		
		2:(*//料框位置抓取*)		
		IF ii=129 THEN(*129表示所有有问题的都抓完了*)
			m_iStep:=4;
		ELSIF ii>0 AND ii<129 AND m_iCheck<>0 
					AND NOT FanucRobotIO.i_xBatteryDetect[0]
					AND NOT FanucRobotIO.i_xBatteryDetect[1]
					AND NOT FanucRobotIO.i_xBatteryDetect[2]
					AND NOT FanucRobotIO.i_xBatteryDetect[3](*4个电池位没料*)
					 (*有不良品*)THEN
			FanucRobotIO.o_xSortStart:=1;(*//从料框取料*)
			FanucRobotIO.o_xColumn[3]:=m_iCoordinateX/8=1;(*XY的偏移量计算在末尾*)
			FanucRobotIO.o_xColumn[2]:=(m_iCoordinateX MOD 8)/4=1;
			FanucRobotIO.o_xColumn[1]:=(m_iCoordinateX MOD 4)/2=1;
			FanucRobotIO.o_xColumn[0]:=(m_iCoordinateX MOD 2)/1=1;
			FanucRobotIO.o_xRow[3]:=m_iCoordinateY/8=1;			
			FanucRobotIO.o_xRow[2]:=(m_iCoordinateY MOD 8)/4=1;
			FanucRobotIO.o_xRow[1]:=(m_iCoordinateY MOD 4)/2=1;
			FanucRobotIO.o_xRow[0]:=(m_iCoordinateY MOD 2)/1=1;
			CASE SortCommunicationIO.i_arriBatteryStatus[ii] OF
			0:(*0表示OCV2的不良品，视为阻值错误处理*)
					FanucRobotIO.o_xPutNumber[1]:=1;					
			1:(*合格*)
					;
			2:(*容量不足*)
					FanucRobotIO.o_xPutNumber[0]:=1;	
			3:(*电压不足*)
					FanucRobotIO.o_xPutNumber[1]:=1;	
			4:(*阻值错误*)
					FanucRobotIO.o_xPutNumber[2]:=1;	
			5:(*电压过高*)
					FanucRobotIO.o_xPutNumber[3]:=1;	
			END_CASE;
		END_IF;
		IF FanucRobotIO.i_xPickOver THEN(*//抓取动作完成*)
			m_iStep:=3;
		END_IF;
	
		3:(*//放入下料皮带线*)
			FanucRobotIO.o_xSortStart:=0;(*//从料框取料*)
			FanucRobotIO.o_xColumn[3]:=0;(*XY的偏移量计算在末尾*)
			FanucRobotIO.o_xColumn[2]:=0;
			FanucRobotIO.o_xColumn[1]:=0;
			FanucRobotIO.o_xColumn[0]:=0;
			FanucRobotIO.o_xRow[3]:=0;
			FanucRobotIO.o_xRow[2]:=0;
			FanucRobotIO.o_xRow[1]:=0;
			FanucRobotIO.o_xRow[0]:=0;	
		IF FanucRobotIO.i_xPutOver THEN(*//抓取动作完成*)
			(*这个得放货完成在复位，方便step2给*)
			FanucRobotIO.o_xPutNumber[0]:=0;
			FanucRobotIO.o_xPutNumber[1]:=0;
			FanucRobotIO.o_xPutNumber[2]:=0;
			FanucRobotIO.o_xPutNumber[3]:=0;
		END_IF;
		m_TONPutover(IN:= FanucRobotIO.o_xPutNumber[0]=0
												AND FanucRobotIO.o_xPutNumber[1]=0
												AND FanucRobotIO.o_xPutNumber[2]=0
												AND FanucRobotIO.o_xPutNumber[3]=0,
			PT:=t#100ms ,Q:= m_xPutover,ET:=m_tPutover );	
			IF LDp(TRUE,m_xPutover)  THEN
				m_iStep:=2;
			END_IF;

		
		4:
		(*4复位所有数据*)
			FanucRobotIO.o_xSortStart:=0;(*//从料框取料*)
			FanucRobotIO.o_xColumn[3]:=0;(*XY的偏移量计算在末尾*)
			FanucRobotIO.o_xColumn[2]:=0;
			FanucRobotIO.o_xColumn[1]:=0;
			FanucRobotIO.o_xColumn[0]:=0;
			FanucRobotIO.o_xRow[3]:=0;
			FanucRobotIO.o_xRow[2]:=0;
			FanucRobotIO.o_xRow[1]:=0;
			FanucRobotIO.o_xRow[0]:=0;	
			FanucRobotIO.o_xPutNumber[0]:=0;
			FanucRobotIO.o_xPutNumber[1]:=0;
			FanucRobotIO.o_xPutNumber[2]:=0;
			FanucRobotIO.o_xPutNumber[3]:=0;

		IF  NOT SortCommunicationIO.o_xSortDone  THEN(*这里表示只给一下2*)
				SortCommunicationIO.o_iSortDonePLCPC:=2;
				SortCommunicationIO.o_xSortDone:=1;
		END_IF;		
		IF SortCommunicationIO.i_iSortDoneAknPCPLC =2 THEN
			SortCommunicationIO.o_iSortDonePLCPC:=1;
			m_iCoordinateX:=1;
			m_iCoordinateY:=1;
		END_IF;
	END_CASE;			
		IF ConveyorIO.xEmpty THEN
				m_iStep:=0;
		END_IF;

	m_iCheck:=	SortCommunicationIO.i_arriBatteryStatus[5]+
							SortCommunicationIO.i_arriBatteryStatus[1]+
							SortCommunicationIO.i_arriBatteryStatus[2]+
							SortCommunicationIO.i_arriBatteryStatus[3]+
							SortCommunicationIO.i_arriBatteryStatus[4];(*连续5个电池都是0，说明这框电池没数据，就不分拣*)
	IF LDP(TRUE,m_iStep=2 AND SortCommunicationIO.i_iInfoWriteDone=2 AND m_iCheck<>0) THEN(*判断哪个地方是有问题的*)
		FOR ii:=ii+1 TO 128 BY 1 DO
			IF SortCommunicationIO.i_arriBatteryStatus[ii]<>1 AND SortCommunicationIO.i_arriBatteryStatus[ii]<>5THEN
				m_iCoordinateX:=((ii-1)/ROW_NUB);
				m_iCoordinateY:=2*((ii-1)MOD ROW_NUB)+((m_iCoordinateX+1) MOD 2);(*把上位机给的编号值对应到二维的偏移上*)(*后面这个意思奇数排+1，偶数排不加*)
				EXIT;
			END_IF;
		END_FOR;
	END_IF;
END_IF;(*g_xauto*)	
IF  g_diDeviceIDSelect=ConveyorIO.diDeviceID AND g_xResetSingle THEN(*复位线体时，同时复位步数和请求，重新来一遍*)
	m_iStep:=0;
END_IF;	
IF  NOT g_xAuto THEN
		SortCommunicationIO.o_iRequestPLCPC:=0;
		SortCommunicationIO.o_iSortDonePLCPC:=0;
END_IF;
END_FUNCTION_BLOCK

PROGRAM START
IF g_xReset THEN
	SM50:=1;
	ELSE
	SM50:=0;
END_IF;
CASE g_iState OF
	0: (*手动*)
	g_xManual:=1;
	g_xAuto:=0;	
	g_xStackLampAmber:=1;
	g_xStackLampGreen:=0;
	g_xRemoteAuto:=0;
	g_xAutoLamp:=0;
	1:(*自动*)
	g_xManual:=0;
	g_xAuto:=1;
	g_xStackLampGreen:=1;
	g_xStackLampAmber:=0;
	g_xRemoteAuto:=0;
	g_xAutoLamp:=1;
	2:	(*远程自动*)
	g_xRemoteAuto:=1;
	g_xStackLampGreen:=1;
	g_xStackLampAmber:=0;
	g_xAuto:=0;
	g_xManual:=0;
	g_xAutoLamp:=0;
	3:(*自动未启动*)
	g_xRemoteAuto:=1;
	g_xStackLampGreen:=SM412;
	g_xStackLampAmber:=0;
	g_xAuto:=0;
	g_xManual:=0;	
	g_xAutoLamp:=0;
END_CASE;

IF g_xAutoSwitch AND g_xAutoStart  THEN  
	g_iState:=1;
END_IF;

IF g_xAutoSwitch AND (g_iState<>1 OR NOT g_xStop)  THEN  
	g_iState:=3;
END_IF;

g_xStackLampRed:=g_xAlarm AND SM412;
g_xBuzzer:=g_xAlarm AND SM412 AND NOT g_xMute;

IF LDF(TRUE,g_xAlarm) THEN
	g_xMute:=0;
END_IF;

IF NOT g_xAutoSwitch  OR g_xEStop=0 THEN 
	g_iState:=0;
END_IF;
IF g_xRemoteAutoStart THEN
	g_iState:=2;
END_IF;
IF g_xPause AND SM412 THEN
	g_xStackLampGreen:=0;
	g_xStackLampAmber:=0;
END_IF;
END_PROGRAM

FUNCTION_BLOCK Switch
VAR_IN_OUT
  ConveyorEntryIO : ConveyorIO;
  ConveyorExitIO : ConveyorIO;
END_VAR
VAR
  m_tonLiftCylinderDelay : TON;  (* 顶升延时 *)
  m_xLiftCylinderDelay : BOOL;
  m_tLiftCylinderDelay : TIME;
  m_tonExitBarDelay : TON;  (* 退出阻挡器延时 *)
  m_tExitBarDelay : TIME;
  m_xExitBarDelay : BOOL;
END_VAR
VAR_IN_OUT
  SwitchIO : SwitchIO;
END_VAR
VAR
  iStep : INT;
  m_xInitial : BOOL;
  m_tonCylinderOvertime : TON;  (* 气缸超时报警定时器 *)
  m_tCylinderOvertimeCurrent : TIME;
END_VAR
(**************************************************
//顶升移载模块，抽象为一条输入输线 ，一条输出输送线
//一个进入阻挡器，一个放出阻挡器，和一个顶升气缸的控制
//程序思路比较混乱，接口不清晰，需要整改
//直接放行的时候有问题
//switchEnable =0的时候   离开线体的PutInto有问题
//增加xPutInto程序
//12-17日   V1.0
//***************************************************)
(*ConveyorEntry(ConveyorMotor:=ConveyorEntryIO);
(*ConveyorExit(ConveyorMotor:=ConveyorExitIO);*)


IF NOT m_xInitial THEN
	SwitchIO.tSetOvertime:=T#5s;
	SwitchIO.xExitEnable:=1;
	m_xInitial:=1;
END_IF;
IF g_xAuto THEN
	CASE iStep OF
		0:(*初始化*)
		ConveyorEntryIO.xLoad:=0;
		ConveyorEntryIO.xUnload:=0;
		ConveyorEntryIO.xPutInto:=0;
		ConveyorExitIO.xLoad:=0;
		ConveyorExitIo.xUnload:=0;
		ConveyorExitIO.xPutInto:=0;
		SwitchIO.xEntryBarCylinderRetract:=0;
		SwitchIO.xExitBarCylinderRetract:=0;
		IF SwitchIO.xLiftCylinderExtendInit THEN
			SwitchIO.xLiftCylinderExtend:=1;
			SwitchIO.xLiftCylinderRetract:=0;
		    IF SwitchIO.xLiftCylinderExtendDetect THEN
			    iStep:=1;
			END_IF; 
			ELSE
			SwitchIO.xLiftCylinderExtend:=0;
			SwitchIO.xLiftCylinderRetract:=1;	
		    IF SwitchIO.xLiftCylinderRetractDetect THEN
			    iStep:=1;
		    END_IF;		
		END_IF;
		1:(*上料*)
        IF SwitchIO.xEntryEnable AND ConveyorEntryIO.xEmpty AND ConveyorExitIO.xEmpty THEN
        	SwitchIO.xEntryBarCylinderRetract:=1;
        	ConveyorEntryIO.xLoad:=1;
        END_IF;
        IF ConveyorEntryIO.xEmpty=0 THEN
        	SwitchIO.xEntryBarCylinderRetract:=0;
        	ConveyorEntryIO.xLoad:=0;
        	ConveyorExitIO.xPutInto:=1;
        END_IF;
        IF m_xLiftCylinderDelay AND  SwitchIO.xSwithEnable AND SwitchIO.xExitEnable THEN
			iStep:=2;
        END_IF;
        IF SwitchIO.xSwithEnable=0 AND m_xLiftCylinderDelay AND SwitchIO.xExitEnable  THEN
			iStep:=3;
        END_IF;
		2:(*顶升*)
		ConveyorExitIO.iProductCategory:=ConveyorEntryIO.iProductCategory;
		ConveyorExitIO.iTaskID:=ConveyorEntryIO.iTaskID;
		ConveyorExitIO.diDesConveyor:=ConveyorEntryIO.diDesConveyor;
		SwitchIO.xExitBarCylinderRetract:=0;
		IF SwitchIO.xLiftCylinderExtendInit THEN
			SwitchIO.xLiftCylinderExtend:=0;
			SwitchIO.xLiftCylinderRetract:=1;
		    ELSE
			SwitchIO.xLiftCylinderExtend:=1;
			SwitchIO.xLiftCylinderRetract:=0;			
		END_IF;

		IF SwitchIO.xLiftCylinderExtendInit THEN
		  	IF SwitchIO.xLiftCylinderRetractDetect THEN
		  		iStep:=4;
		  	END_IF;
		  	ELSE
		  	IF SwitchIO.xLiftCylinderExtendDetect THEN
				iStep:=4; 
		  	END_IF;
		END_IF;
		3:(*放行*)	
		ConveyorExitIO.iProductCategory:=ConveyorEntryIO.iProductCategory;
		ConveyorExitIO.iTaskID:=ConveyorEntryIO.iTaskID;
		ConveyorExitIO.diDesConveyor:=ConveyorEntryIO.diDesConveyor;
		SwitchIO.xExitBarCylinderRetract:=1;
		ConveyorExitIO.xPutInto:=0;
		iStep:=4;
		4:(*下料*)
		(*通过出料传输线下料*)
		IF SwitchIO.xExitEnable  AND m_xExitBarDelay AND NOT SwitchIO.xExitBarCylinderRetract  THEN		  
		  	ConveyorExitIO.xUnload:=1;
			ELSE
		  	ConveyorExitIO.xUnload:=0;
		END_IF;	
		(*通过进料传输线下料*)
		IF SwitchIO.xExitEnable  AND m_xExitBarDelay  AND SwitchIO.xExitBarCylinderRetract THEN		  
		  	ConveyorEntryIO.xUnload:=1;
			ELSE
		  	ConveyorEntryIO.xUnload:=0;
		END_IF;			    	
		IF (ConveyorExitIO.xEmpty OR ConveyorEntryIO.xEmpty) AND m_xExitBarDelay  THEN
		  	ConveyorExitIO.xPutInto:=1;
		  	ConveyorEntryIO.xPutInto:=1;
			iStep:=0; 
		END_IF;
	END_CASE;
	m_tonLiftCylinderDelay(IN:=NOT ConveyorEntryIO.xEmpty AND iStep=1 ,PT:= T#1S ,Q:= m_xLiftCylinderDelay ,ET:=m_tLiftCylinderDelay );
	m_tonExitBarDelay(IN:=iStep=4 ,PT:= T#1s ,Q:= m_xExitBarDelay ,ET:= m_tExitBarDelay);
END_IF;
(*复位程序*)
IF (g_xResetSingle AND  (g_diDeviceIDSelect=ConveyorEntryIO.diDeviceID OR g_diDeviceIDSelect=ConveyorExitIO.diDeviceID))
	OR LDP(TRUE,SwitchIO.xLiftCylinderExtendInit) 
	OR LDF(TRUE,SwitchIO.xLiftCylinderExtendInit) 
	OR LDP(TRUE,SwitchIO.xPutInto)  THEN
	ConveyorEntryIO.xPutInto:=1;
	ConveyorExitIO.xPutInto:=1;
	iStep:=0;
END_IF;

IF g_xManual  THEN
	iStep:=0;
	ConveyorEntryIO.xLoad:=0;
    ConveyorEntryIO.xUnload:=0;
	ConveyorEntryIO.xPutInto:=0;
	ConveyorExitIO.xLoad:=0;
	ConveyorExitIo.xUnload:=0;
	ConveyorExitIO.xPutInto:=0;
	SwitchIO.xEntryBarCylinderRetract:=0;
	SwitchIO.xExitBarCylinderRetract:=0;
	IF SwitchIO.xEntryBarCylinderRetractButton THEN
		SwitchIO.xEntryBarCylinderRetract:=1;
		ELSE
		SwitchIO.xEntryBarCylinderRetract:=0;
	END_IF;
	IF SwitchIO.xExitBarCylinderRetractButton THEN
		SwitchIO.xExitBarCylinderRetract:=1;
		ELSE
		SwitchIO.xExitBarCylinderRetract:=0;
	END_IF;
	IF SwitchIO.xLiftCylinderExtendButton AND NOT SwitchIO.xLiftCylinderRetractButton THEN
		SwitchIO.xLiftCylinderExtend:=1;
		SwitchIO.xLiftCylinderRetract:=0;
	END_IF;
	IF NOT SwitchIO.xLiftCylinderExtendButton AND  SwitchIO.xLiftCylinderRetractButton THEN
		SwitchIO.xLiftCylinderExtend:=0;
		SwitchIO.xLiftCylinderRetract:=1;
	END_IF;		 
END_IF;
(*气缸超时报警*)
m_tonCylinderOvertime(IN:= (SwitchIO.xLiftCylinderExtend AND NOT SwitchIO.xLiftCylinderExtendDetect) 
OR  (SwitchIO.xLiftCylinderRetract AND NOT SwitchIO.xLiftCylinderRetractDetect) ,
PT:= SwitchIO.tSetOvertime ,Q:= SwitchIO.xOvertimeAlarm ,ET:= m_tCylinderOvertimeCurrent );
END_FUNCTION_BLOCK

PROGRAM TCP
VAR
  m_ton1ReceiveHeartbeat : TON;
  m_t1RecHeartbeatCurrentTime : TIME;
  m_tonAutoClose : TON;
  m_xAutoClose : BOOL;
  m_tAutoCloseCurrentTime : TIME;
  m_tonReconnect : TON;
  m_xReconnect : BOOL;
  m_tReconnectCurrentTime : TIME;
  m_ton5ReceiveHeartbeat : TON;
  m_t5RecHeartbeatCurrentTime : TIME;
  m_ton2ReceiveHeartbeat : TON;
  m_t2RecHeartbeatCurrentTime : TIME;
END_VAR
(*与RGV通信*)
D200:=18;
(*m_tonReconnect(IN:= NOT SD1282.0 AND NOT SD1284.0,PT:=T#5s  ,Q:=m_xReconnect ,ET:=m_tReconnectCurrentTime);*)
(*1282打开完成状态*)(*1284打开请求状态*)
(*SP_SOCOPEN(m_xReconnect  AND SD1288.A , "U0", K1 , D110 , M100);*)
(*1288.A设备连接状态*)
SP_SOCSND( SM412 AND SD1282.5 , "U0" , K6 , D100, D200, M102 );
SP_SOCRCV( SD1282.5 AND SD1286.5 AND NOT M104 , "U0" , K6, D300 , D400 ,M104 );
(*1286数据接收状态*)
(*m_tonAutoClose(IN:= SD1284.0 AND NOT SD1282.0 ,PT:=T#5s,Q:=m_xAutoClose ,ET:= m_tAutoCloseCurrentTime );
SP_SOCCLOSE( LDF(TRUE,SD1282.0) OR m_xAutoClose  , "U0" , K1, D120, M106 );*)
D203.F:=SM413;
m_ton1ReceiveHeartbeat(IN:=NOT LDP(TRUE, D403.F) ,PT:= t#5S ,Q:= g_xRGVTcpFailed ,ET:= m_t1RecHeartbeatCurrentTime);
IF g_xRGVTcpFailed THEN
	M104:=SM413;(*通讯失败有可能是接收模块没动作，重启接收模块*)
	D400:=0;
	D401:=0;
END_IF;



(*与40通信*)
D220:=2;
(*m_tonReconnect(IN:= NOT SD1282.0 AND NOT SD1284.0,PT:=T#5s  ,Q:=m_xReconnect ,ET:=m_tReconnectCurrentTime);*)
(*1282打开完成状态*)(*1284打开请求状态*)
(*SP_SOCOPEN(m_xReconnect  AND SD1288.A , "U0", K1 , D110 , M100);*)
(*1288.A设备连接状态*)
SP_SOCSND( SM412 AND SD1282.4 , "U0" , K5, D120, D220, M122 );
SP_SOCRCV( SD1282.4 AND SD1286.4 AND NOT M124 , "U0" , K5, D320 , D420 ,M124 );
(*1286数据接收状态*)
(*m_tonAutoClose(IN:= SD1284.0 AND NOT SD1282.0 ,PT:=T#5s,Q:=m_xAutoClose ,ET:= m_tAutoCloseCurrentTime );
SP_SOCCLOSE( LDF(TRUE,SD1282.0) OR m_xAutoClose  , "U0" , K1, D120, M106 );*)
D221.F:=SM413;
m_ton2ReceiveHeartbeat(IN:=NOT LDP(TRUE, D421.F) ,PT:= t#5S ,Q:= g_x60TcpFailed ,ET:= m_t2RecHeartbeatCurrentTime);
IF g_x60TcpFailed THEN
	M124:=SM413;(*通讯失败有可能是接收模块没动作，重启接收模块*)
	D420:=0;
	D421:=0;
END_IF;
END_PROGRAM

FUNCTION_BLOCK UConveyor
VAR
  iStep : INT;
END_VAR
VAR_IN_OUT
  ConveyorIOLeft : ConveyorIO;  (* U的左半边 *)
  ConveyorIORight : ConveyorIO;  (* U的右半边 *)
  ConveyorIODown : ConveyorIO;  (* U的下边一横 *)
  UConveyorIO : UConveyorIO;  (* 顶升,阻挡 *)
END_VAR
VAR
  m_xInitial : BOOL;
  m_tonCylinderOvertime : TON;  (* 气缸超时报警定时器 *)
  m_tCylinderOvertimeCurrent : TIME;
  m_tonExitBarDelay : TON;  (* 退出阻挡器延时 *)
  m_tExitBarDelay : TIME;
  m_xExitBarDelay : BOOL;
  m_TonStep0 : TON;  (* Step为0延时 *)
  m_xStep0 : BOOL;  (* Step为0延时 *)
  m_tStep0 : TIME;  (* Step为0延时 *)
END_VAR
(*                                                                                                          
初始化中增加气缸复位，气缸位置有BUG
//*)
IF NOT m_xInitial THEN
	UConveyorIO.tSetOvertime:=T#5s;
	UConveyorIO.xExitEnable1:=1;
	UConveyorIO.xExitEnable2:=1;
	UConveyorIO.xExitEnable3:=1;
	m_xInitial:=1;
END_IF;
(*外部不用写ConveyorDown的开关，会自己根据来料的产品信息判断停哪个光电*)
IF UConveyorIO.iTask=1 AND ConveyorIODown.diDesConveyorIn=ConveyorIOLeft.diDeviceID THEN
	ConveyorIODown.xCWPresent:=ConveyorIOLeft.xCCWPresent;
ELSIF UConveyorIO.iTask=1 AND ConveyorIODown.diDesConveyorIn=ConveyorIORight.diDeviceID THEN
	ConveyorIODown.xCWPresent:=ConveyorIORight.xCCWPresent;
ELSE
	ConveyorIODown.xCWPresent:=ConveyorIOLeft.xCCWPresent OR ConveyorIORight.xCCWPresent;
END_IF;
(*这里判断什么时候直接放行，左右都不需要，也不是0，就放走*)
IF  NOT(ConveyorIODown.diDesConveyor=ConveyorIOLeft.diDeviceID 
		OR  ConveyorIODown.diDesConveyor=ConveyorIORight.diDeviceID 
		OR ConveyorIODown.diDesConveyor=0) THEN
	UConveyorIO.xPassEnable:=1;
ELSE
	UConveyorIO.xPassEnable:=0;
END_IF;	
IF g_xAuto THEN	
(*	//加个Step为0的延时，防止扫描周期的影响*)
	m_TonStep0(IN:= iStep=0 ,PT:= t#100ms ,Q:= m_xStep0 ,ET:= m_tStep0 );
	(*//这个是留给阻挡动作的时间*)
	m_tonExitBarDelay(IN:=iStep=4 ,PT:= T#1s ,Q:= m_xExitBarDelay ,ET:= m_tExitBarDelay);
CASE UConveyorIO.iTask OF(*这个Task做抢占，可做LastTask保护*)
0:(*各种初始化，能自动去3*)
	ConveyorIODown.xLoad:=0;
	ConveyorIOleft.xLoad:=0;
	ConveyorIORight.xLoad:=0;
	ConveyorIODown.xUnload:=0;
	ConveyorIOLeft.xUnload:=0;
	ConveyorIORight.xUnload:=0;
	ConveyorIODown.xPutInto:=0;
	ConveyorIOLeft.xPutInto:=0;
	ConveyorIORight.xPutInto:=0;	
	UConveyorIO.xExitBarCylinderRetract1:=0;
	UConveyorIO.xExitBarCylinderRetract2:=0;	
	UConveyorIO.xLiftCylinderRetract1:=1;
	UConveyorIO.xLiftCylinderRetract2:=1;
	UConveyorIO.xLiftCylinderExtend1:=0;
	UConveyorIO.xLiftCylinderExtend2:=0;
1:(*上料*)
	CASE iStep OF
	0:(*各种初始化，能自动去3*)
		ConveyorIODown.xLoad:=0;
		ConveyorIOleft.xLoad:=0;
		ConveyorIORight.xLoad:=0;
		ConveyorIODown.xUnload:=0;
		ConveyorIOLeft.xUnload:=0;
		ConveyorIORight.xUnload:=0;
		UConveyorIO.xExitBarCylinderRetract1:=0;
		UConveyorIO.xExitBarCylinderRetract2:=0;
		UConveyorIO.xBatteryError:=0;
		ConveyorIODown.xPutInto:=0;
		ConveyorIOLeft.xPutInto:=0;
		ConveyorIORight.xPutInto:=0;	
	(*	//根据是否有料判断去1还是3，但会等一个延时*)
		IF m_xStep0 AND  ConveyorIODown.xEmpty THEN
			iStep:=1;
		ELSIF m_xStep0 AND NOT ConveyorIODown.xEmpty THEN
			iStep:=3;
		END_IF;	
	1:(*顶升初始化，等load*)
		(*//左顶升*)
		IF UConveyorIO.xLiftCylinderExtendInit1 THEN
			UConveyorIO.xLiftCylinderExtend1:=1;
			UConveyorIO.xLiftCylinderRetract1:=0;
		ELSE
			UConveyorIO.xLiftCylinderExtend1:=0;
			UConveyorIO.xLiftCylinderRetract1:=1;
		END_IF;
	(*	//右顶升*)
		IF UConveyorIO.xLiftCylinderExtendInit2 THEN
			UConveyorIO.xLiftCylinderExtend2:=1;
			UConveyorIO.xLiftCylinderRetract2:=0;
			ELSE
			UConveyorIO.xLiftCylinderExtend2:=0;
			UConveyorIO.xLiftCylinderRetract2:=1;
		END_IF;
		(*//顶升到位，等上料信号*)
		IF 	((UConveyorIO.xLiftCylinderExtendInit1 AND UConveyorIO.xLiftCylinderExtendDetect1)
				OR (NOT UConveyorIO.xLiftCylinderExtendInit1 AND UConveyorIO.xLiftCylinderRetractDetect1))
			AND	((UConveyorIO.xLiftCylinderExtendInit2 AND UConveyorIO.xLiftCylinderExtendDetect2)
		   		OR (NOT UConveyorIO.xLiftCylinderExtendInit2 AND UConveyorIO.xLiftCylinderRetractDetect2))		
			AND	UConveyorIO.xEntryEnable1 THEN(*有上料请求1*)
		   	ConveyorIODown.xLoad:=1;
			iStep:=2;
		END_IF;
	2:(*Load完成*)
		(*去右臂时才需要阻挡1放行,其他情况阻挡1挡住*)
		UConveyorIO.xExitBarCylinderRetract1:=ConveyorIODown.diDesConveyorIn=ConveyorIORight.diDeviceID;
		IF NOT ConveyorIODown.xEmpty THEN
			ConveyorIODown.xLoad:=0;
			ConveyorIOLeft.xPutInto:=1;
			ConveyorIOright.xPutInto:=1;
			istep:=3;
		END_IF;
	3:(*顶升等Unload，这里等有了ExitEnable再顶升，因为可能有地方需要允许了再升降，比如倍速链*)
		(*//电池检测保护，防止把带电池的料框送进去了*)
		IF (ConveyorIODown.diDesConveyor=ConveyorIOLeft.diDeviceID OR ConveyorIODown.diDesConveyor=ConveyorIORight.diDeviceID)
			AND	(UConveyorIO.xBatteryDetect1 OR UConveyorIO.xBatteryDetect2)(*在下面时检测*)
			AND UConveyorIO.xLiftCylinderRetractDetect1 AND UConveyorIO.xLiftCylinderRetractDetect2 THEN
			UConveyorIO.xBatteryError:=1;
		END_IF;	
		(*//左侧顶升控制*)
		IF (ConveyorIODown.diDesConveyor=ConveyorIOLeft.diDeviceID AND UConveyorIO.xExitEnable2 AND NOT UConveyorIO.xBatteryError)THEN
			IF UConveyorIO.xLiftCylinderExtendInit1 THEN
				UConveyorIO.xLiftCylinderExtend1:=0;
				UConveyorIO.xLiftCylinderRetract1:=1;
			ELSE
				UConveyorIO.xLiftCylinderExtend1:=1;
				UConveyorIO.xLiftCylinderRetract1:=0;
			END_IF;
			IF(NOT UConveyorIO.xLiftCylinderExtendInit1 AND UConveyorIO.xLiftCylinderExtendDetect1)
				OR (UConveyorIO.xLiftCylinderExtendInit1 AND UConveyorIO.xLiftCylinderRetractDetect1)THEN
				ConveyorIOLeft.xPutInto:=0;
				ConveyorIOright.xPutInto:=0;
				iStep:=4;
			END_IF;
		END_IF;	
		(*//右侧顶升控制*)
		IF (ConveyorIODown.diDesConveyor=ConveyorIORight.diDeviceID AND UConveyorIO.xExitEnable3 AND NOT UConveyorIO.xBatteryError)THEN
			IF UConveyorIO.xLiftCylinderExtendInit2 THEN
				UConveyorIO.xLiftCylinderExtend2:=0;
				UConveyorIO.xLiftCylinderRetract2:=1;
			ELSE
				UConveyorIO.xLiftCylinderExtend2:=1;
				UConveyorIO.xLiftCylinderRetract2:=0;
			END_IF;
			IF(NOT UConveyorIO.xLiftCylinderExtendInit2 AND UConveyorIO.xLiftCylinderExtendDetect2)
				OR (UConveyorIO.xLiftCylinderExtendInit2 AND UConveyorIO.xLiftCylinderRetractDetect2) THEN
				ConveyorIOLeft.xPutInto:=0;
				ConveyorIOright.xPutInto:=0;
				iStep:=4;
			END_IF;
		END_IF;	
	(*	//直接放行控制*)
		IF UConveyorIO.xPassEnable AND UConveyorIO.xExitEnable1 AND NOT UConveyorIO.xBatteryError THEN
			IF UConveyorIO.xLiftCylinderExtendInit1 THEN
				UConveyorIO.xLiftCylinderExtend1:=1;
				UConveyorIO.xLiftCylinderRetract1:=0;
			ELSE
				UConveyorIO.xLiftCylinderExtend1:=0;
				UConveyorIO.xLiftCylinderRetract1:=1;
			END_IF;
			IF UConveyorIO.xLiftCylinderExtendInit2 THEN
				UConveyorIO.xLiftCylinderExtend2:=1;
				UConveyorIO.xLiftCylinderRetract2:=0;
			ELSE
				UConveyorIO.xLiftCylinderExtend2:=0;
				UConveyorIO.xLiftCylinderRetract2:=1;
			END_IF;
			IF((UConveyorIO.xLiftCylinderExtendInit1 AND UConveyorIO.xLiftCylinderExtendDetect1)
 OR (NOT UConveyorIO.xLiftCylinderExtendInit1 AND UConveyorIO.xLiftCylinderRetractDetect1))
				AND((UConveyorIO.xLiftCylinderExtendInit2 AND UConveyorIO.xLiftCylinderExtendDetect2)
 OR (NOT UConveyorIO.xLiftCylinderExtendInit2 AND UConveyorIO.xLiftCylinderRetractDetect2))THEN
				UConveyorIO.xExitBarCylinderRetract1:=1;
				UConveyorIO.xExitBarCylinderRetract2:=1;
				ConveyorIOLeft.xPutInto:=0;
				ConveyorIOright.xPutInto:=0;
				iStep:=4;
			END_IF;	
		END_IF;
	4:(*Unload完成，回0*)
			IF ConveyorIODown.diDesConveyor=ConveyorIOLeft.diDeviceID AND UConveyorIO.xExitEnable2 AND m_xExitBarDelay THEN
				ConveyorIOLeft.xUnload:=1;
			ELSIF ConveyorIODown.diDesConveyor=ConveyorIORight.diDeviceID AND UConveyorIO.xExitEnable3 AND m_xExitBarDelay THEN
				ConveyorIORight.xUnload:=1;
			ELSIF UConveyorIO.xPassEnable AND UConveyorIO.xExitEnable1 AND m_xExitBarDelay THEN
				ConveyorIODown.xUnload:=1;
			ELSE
				ConveyorIODown.xUnload:=0;
				ConveyorIOLeft.xUnload:=0;
				ConveyorIORight.xUnload:=0;
			END_IF;	
		IF ( (ConveyorIODown.diDesConveyor=ConveyorIOLeft.diDeviceID  AND LDF(TRUE,UConveyorIO.xExitEnable2))
		  OR(ConveyorIODown.diDesConveyor=ConveyorIORight.diDeviceID AND LDF(TRUE,UConveyorIO.xExitEnable3))
		  OR(UConveyorIO.xPassEnable AND LDF(TRUE,UConveyorIO.xExitEnable1)) )AND m_xExitBarDelay  THEN
			ConveyorIODown.xUnload:=0;
			ConveyorIOLeft.xUnload:=0;
			ConveyorIORight.xUnload:=0;
			ConveyorIODown.xPutInto:=1;
			ConveyorIOLeft.xPutInto:=1;
			ConveyorIORight.xPutInto:=1;
			UConveyorIO.xExitBarCylinderRetract1:=0;
			UConveyorIO.xExitBarCylinderRetract2:=0;
			iStep:=0;
		END_IF;
	END_CASE;
2:(*左下料*)
	CASE iStep OF
	0:(*各种初始化，能自动去3*)
		ConveyorIODown.xLoad:=0;
		ConveyorIOleft.xLoad:=0;
		ConveyorIORight.xLoad:=0;
		ConveyorIODown.xUnload:=0;
		ConveyorIOLeft.xUnload:=0;
		ConveyorIORight.xUnload:=0;
		UConveyorIO.xBatteryError:=0;
		UConveyorIO.xExitBarCylinderRetract1:=0;
		UConveyorIO.xExitBarCylinderRetract2:=0;
		ConveyorIODown.xPutInto:=0;
		ConveyorIOLeft.xPutInto:=0;
		ConveyorIORight.xPutInto:=0;
		IF m_xStep0 AND  ConveyorIODown.xEmpty THEN
			iStep:=1;
		ELSIF m_xStep0 AND NOT ConveyorIODown.xEmpty THEN
			iStep:=3;
		END_IF;	
	1:(*左顶升动作，等load*)
		IF UConveyorIO.xLiftCylinderExtendInit1 THEN
			UConveyorIO.xLiftCylinderExtend1:=0;
			UConveyorIO.xLiftCylinderRetract1:=1;
			ELSE
			UConveyorIO.xLiftCylinderExtend1:=1;
			UConveyorIO.xLiftCylinderRetract1:=0;
		END_IF;
		IF ((NOT UConveyorIO.xLiftCylinderExtendInit1 AND UConveyorIO.xLiftCylinderExtendDetect1)
			OR ( UConveyorIO.xLiftCylinderExtendInit1 AND UConveyorIO.xLiftCylinderRetractDetect1))
			AND UConveyorIO.xEntryEnable2 THEN(*有上料请求1*)
		   	ConveyorIOLeft.xLoad:=1;
			iStep:=2;
		END_IF;
	2:(*Load完成*)
		IF NOT ConveyorIOLeft.xEmpty THEN
			ConveyorIOLeft.xLoad:=0;
			ConveyorIODown.xPutInto:=1;
			ConveyorIODown.diDesConveyor:=ConveyorIOLeft.diDesConveyor;
			istep:=3;
		END_IF;
	3:(*顶升等Unload，这里等有了ExitEnable再顶升，因为可能有地方需要允许了再升降，比如倍速链*)
		UConveyorIO.xExitBarCylinderRetract1:=1;
		UConveyorIO.xExitBarCylinderRetract2:=1;
		IF  UConveyorIO.xExitEnable1 THEN
			IF UConveyorIO.xLiftCylinderExtendInit1 THEN
				UConveyorIO.xLiftCylinderExtend1:=1;
				UConveyorIO.xLiftCylinderRetract1:=0;
			ELSE
				UConveyorIO.xLiftCylinderExtend1:=0;
				UConveyorIO.xLiftCylinderRetract1:=1;
			END_IF;
			IF(( UConveyorIO.xLiftCylinderExtendInit1 AND UConveyorIO.xLiftCylinderExtendDetect1)
				OR (NOT UConveyorIO.xLiftCylinderExtendInit1 AND UConveyorIO.xLiftCylinderRetractDetect1))THEN
				ConveyorIODown.xPutInto:=0;
				iStep:=4;
			END_IF;	
		END_IF;
	4:(*Unload完成，回0*)
		IF  UConveyorIO.xExitEnable1 AND m_xExitBarDelay THEN
			ConveyorIODown.xUnload:=1;
		ELSE
			ConveyorIODown.xUnload:=0;
		END_IF;	
		IF NOT UConveyorIO.xExitEnable1 AND m_xExitBarDelay   THEN
			ConveyorIODown.xUnload:=0;
			ConveyorIOLeft.xUnload:=0;
			ConveyorIORight.xUnload:=0;
			ConveyorIODown.xPutInto:=1;
			ConveyorIOLeft.xPutInto:=1;
			ConveyorIORight.xPutInto:=1;
			UConveyorIO.xExitBarCylinderRetract1:=0;
			UConveyorIO.xExitBarCylinderRetract2:=0;
			iStep:=0;
		END_IF;
	END_CASE;
3:(*上料到出口*)
	CASE iStep OF
	0:(*各种初始化，能自动去3*)
		ConveyorIODown.xLoad:=0;
		ConveyorIOleft.xLoad:=0;
		ConveyorIORight.xLoad:=0;
		ConveyorIODown.xUnload:=0;
		ConveyorIOLeft.xUnload:=0;
		ConveyorIORight.xUnload:=0;
		UConveyorIO.xBatteryError:=0;
		UConveyorIO.xExitBarCylinderRetract1:=0;
		UConveyorIO.xExitBarCylinderRetract2:=0;
		ConveyorIODown.xPutInto:=0;
		ConveyorIOLeft.xPutInto:=0;
		ConveyorIORight.xPutInto:=0;
		IF m_xStep0 AND  ConveyorIODown.xEmpty THEN
			iStep:=1;
		ELSIF m_xStep0 AND NOT ConveyorIODown.xEmpty THEN
			iStep:=3;
		END_IF;	
	1:(*右顶升动作，等load*)
		IF UConveyorIO.xLiftCylinderExtendInit2 THEN
			UConveyorIO.xLiftCylinderExtend2:=0;
			UConveyorIO.xLiftCylinderRetract2:=1;
		ELSE
			UConveyorIO.xLiftCylinderExtend2:=1;
			UConveyorIO.xLiftCylinderRetract2:=0;
		END_IF;
		IF ((NOT UConveyorIO.xLiftCylinderExtendInit2 AND UConveyorIO.xLiftCylinderExtendDetect2)
			OR ( UConveyorIO.xLiftCylinderExtendInit2 AND UConveyorIO.xLiftCylinderRetractDetect2))
			AND UConveyorIO.xEntryEnable3 THEN(*有上料请求1*)
		   	ConveyorIORight.xLoad:=1;
			iStep:=2;
		END_IF;
	2:(*Load完成*)
		IF NOT ConveyorIORight.xEmpty THEN
			ConveyorIORight.xLoad:=0;
			ConveyorIODown.diDesConveyor:=ConveyorIORight.diDesConveyor;
			ConveyorIODown.xPutInto:=1;
			istep:=3;
		END_IF;
	3:(*顶升恢复等Unload，这里等有了ExitEnable再顶升，因为可能有地方需要允许了再升降，比如倍速链*)
		UConveyorIO.xExitBarCylinderRetract2:=1;
		IF  UConveyorIO.xExitEnable1 THEN(**)
			IF UConveyorIO.xLiftCylinderExtendInit2 THEN
				UConveyorIO.xLiftCylinderExtend2:=1;
				UConveyorIO.xLiftCylinderRetract2:=0;
			ELSE
				UConveyorIO.xLiftCylinderExtend2:=0;
				UConveyorIO.xLiftCylinderRetract2:=1;
			END_IF;
		END_IF;
		IF UConveyorIO.xExitEnable1 THEN(**)
			IF(( UConveyorIO.xLiftCylinderExtendInit2 AND UConveyorIO.xLiftCylinderExtendDetect2)
				OR (NOT UConveyorIO.xLiftCylinderExtendInit2 AND UConveyorIO.xLiftCylinderRetractDetect2))THEN
				ConveyorIODown.xPutInto:=0;
				iStep:=4;
			END_IF;	
		END_IF;
	4:(*Unload完成，回0*)
		IF  UConveyorIO.xExitEnable1 AND m_xExitBarDelay THEN
			ConveyorIODown.xUnload:=1;
		ELSE
			ConveyorIODown.xUnload:=0;
		END_IF;	
		IF NOT UConveyorIO.xExitEnable1 AND m_xExitBarDelay  THEN
			ConveyorIODown.xUnload:=0;
			ConveyorIOLeft.xUnload:=0;
			ConveyorIORight.xUnload:=0;
			ConveyorIODown.xPutInto:=1;
			ConveyorIOLeft.xPutInto:=1;
			ConveyorIORight.xPutInto:=1;
			UConveyorIO.xExitBarCylinderRetract1:=0;
			UConveyorIO.xExitBarCylinderRetract2:=0;
			iStep:=0;
		END_IF;
	END_CASE;
END_CASE;(*iTask*)
END_IF;(*g_xAuto那个IF*)
(*复位程序*)
IF (g_xResetSingle AND  (g_diDeviceIDSelect=ConveyorIOLeft.diDeviceID 
 	 OR g_diDeviceIDSelect=ConveyorIORight.diDeviceID
 	 OR g_diDeviceIDSelect=ConveyorIODown.diDeviceID))
	OR LDP(TRUE,UConveyorIO.xLiftCylinderExtendInit1) 
	OR LDF(TRUE,UConveyorIO.xLiftCylinderExtendInit1) 
	OR LDP(TRUE,UConveyorIO.xPutInto)  THEN
	ConveyorIODown.xPutInto:=1;
	ConveyorIOLeft.xPutInto:=1;
	ConveyorIORight.xPutInto:=1;
	iStep:=0;
END_IF;
(*手动*)
IF g_xManual  THEN
	iStep:=0;
	ConveyorIODown.xLoad:=0;
	ConveyorIOleft.xLoad:=0;
	ConveyorIORight.xLoad:=0;
	ConveyorIODown.xUnload:=0;
	ConveyorIOLeft.xUnload:=0;
	ConveyorIORight.xUnload:=0;
	ConveyorIODown.xPutInto:=0;
	ConveyorIOLeft.xPutInto:=0;
	ConveyorIORight.xPutInto:=0;
	UConveyorIO.xBatteryError:=0;
	UConveyorIO.xLiftCylinderExtend1:=UConveyorIO.xLiftCylinderExtendButton1 AND NOT UConveyorIO.xLiftCylinderRetractButton1;
	UConveyorIO.xLiftCylinderRetract1:=UConveyorIO.xLiftCylinderRetractButton1 AND NOT UConveyorIO.xLiftCylinderExtendButton1;
	UConveyorIO.xLiftCylinderExtend2:=UConveyorIO.xLiftCylinderExtendButton2 AND NOT UConveyorIO.xLiftCylinderRetractButton2;
	UConveyorIO.xLiftCylinderRetract2:=UConveyorIO.xLiftCylinderRetractButton2 AND NOT UConveyorIO.xLiftCylinderExtendButton2;
	UConveyorIO.xExitBarCylinderRetract1:=UConveyorIO.xExitBarCylinderRetractButton1;
	UConveyorIO.xExitBarCylinderRetract2:=UConveyorIO.xExitBarCylinderRetractButton2;
END_IF;	
(*气缸超时报警*)
m_tonCylinderOvertime(IN:= (UConveyorIO.xLiftCylinderExtend1 AND NOT UConveyorIO.xLiftCylinderExtendDetect1) 
 		OR  (UConveyorIO.xLiftCylinderRetract1 AND NOT UConveyorIO.xLiftCylinderRetractDetect1)
 		OR	(UConveyorIO.xLiftCylinderExtend2 AND NOT UConveyorIO.xLiftCylinderExtendDetect2) 
 		OR  (UConveyorIO.xLiftCylinderRetract2 AND NOT UConveyorIO.xLiftCylinderRetractDetect2),
 PT:= UConveyorIO.tSetOvertime ,Q:=UConveyorIO.xOvertimeAlarm ,ET:=m_tCylinderOvertimeCurrent );
END_FUNCTION_BLOCK

PROGRAM 复制

END_PROGRAM
